
   hm  24. oct 2007        rev 1.4
       changed dst calculation because function dst was upgraded no error in DCF77 only a change in DST

   hm  12. nov 2007        rev 1.5
       changed time_offset from time to integer to allow for negative offset time zones

   hm  8. dec 2007     rev 1.6
       corrected an error in time_zone calculation

   hm 23. jan 2008     rev 1.7
       added sdt input which is used to initialize rtc and rtc1 during first cycle.

   hm 16. mar 2008     rev 1.8
       changed output weekday to wday and dst to ds for compatibility reasons

   hm  19. apr. 2008   rev 1.9
       added input dsi to allow to set daylight savings time when SDT is TRUE.
       added asynchronous SET input

   hm  7. oct. 2008    rev 1.10
       changed function weekday to day_of_week

   *)
END_FUNCTION_BLOCK

FUNCTION_BLOCK "HOLIDAY"   // FB28, SCL
TITLE = HOLIDAY
{ S7_Optimized_Access := 'FALSE' }
AUTHOR : hugo
FAMILY : TIDT
NAME : HOLIDAY
VERSION : 2.0
// holiday calculates if a given day is a holiday and displays the name of the holiday as string as well as a boolean flag to indicate a holiday.
// the holidays are specified in the country setup under global constants.
// a holiday can be of fixed date for example new years day on january 1st.
// a holiday can have a fixed offset from easter sunday as for most church holidays.
// a holiday can be a specific weekday before a fixed date, for example buss und bettag is the last wednesday before nov 23rd.
// with a simple f_use flag any specific holiday can be turned on or off if needed.
// 
// uses: LOCATION (DB5)
//       HOLIDAY_DATA (UDT9)
//       YEAR_OF_DATE (FC219)
//       EASTER (FC186)
//       SET_DATE (FC213)
//       LEAP_YEAR (FC194)
//       DAY_OF_WEEK (FC179)
//       DATE_ADD (FC176)
//       MONTH_OF_DATE (FC202)
//       DAY_OF_YEAR (FC180)
//       DATE_DINT (FC405)
//       LEAP_OF_DATE (FC193)
//       DAY_OF_MONTH (FC178)
   VAR_INPUT
      DATE_IN : Date;
      LANGU : Int;
      FRIDAY : Bool;
      SATURDAY : Bool;
      SUNDAY : Bool;
      SIZE : Int := 29;
   END_VAR
   VAR_OUTPUT
      Y : Bool;
      _NAME : String[30];
   END_VAR
   VAR_IN_OUT
      HOLIDAYS : Array[0..29] of "HOLIDAY_DATA";
   END_VAR
   VAR
      last_active : Date;
      ostern : Date;
      i : Int;
      jahr : Int;
      x_date : Date;
      lx : Int;
      wdx : Int;
   END_VAR
BEGIN


   (* for performance reasons only activate once a day *)
   IF #last_active = #DATE_IN THEN RETURN; END_IF;
   #last_active := #DATE_IN;

   (* determine language *)
   IF #LANGU = 0 THEN
     #lx := "LANGUAGE".DEFAULT;
   ELSE
     #lx := MIN(IN1:="LANGUAGE".LMAX,IN2:=#LANGU);
   END_IF;

   (* berechnung von ostern für das aktuelle jahr *)
   #jahr := "YEAR_OF_DATE"(#DATE_IN);
   #ostern := "EASTER"(#jahr);
   #wdx := "DAY_OF_WEEK"(#DATE_IN);
   #Y := FALSE;

   (* check for holidays *)
   FOR #i := 0 TO #SIZE DO
     #x_date := "SET_DATE"(YEAR:=#jahr, MONTH:=#HOLIDAYS[#i].MONTH , DAY:=#HOLIDAYS[#i].DAY);
     IF #HOLIDAYS[#i].USE = 1 AND #HOLIDAYS[#i].MONTH > 0 THEN
       (* check for fixed date holiday *)
       IF #x_date = #DATE_IN THEN
         #Y := TRUE;
         #_NAME := #HOLIDAYS[#i]BLKMOV_NAME;
         RETURN;
       END_IF;
     ELSIF #HOLIDAYS[#i].USE = 1 AND #HOLIDAYS[#i].MONTH = 0 THEN
       (* check for holiday in reference to easter *)
       IF "DATE_ADD"(IDATE:=#ostern, D:=#HOLIDAYS[#i].DAY ,W:=0,M:=0,Y:=0) = #DATE_IN THEN
         #Y := TRUE;
         #_NAME := #HOLIDAYS[#i]._NAME;
         RETURN;
       END_IF;
     ELSIF #HOLIDAYS[#i].USE < 0 THEN
       (* check for holiday on a weekday before date *)
       IF "DAY_OF_WEEK"(#DATE_IN) = ABS(#HOLIDAYS[#i].USE) AND #DATE_IN < #x_date AND #DATE_IN >= "DATE_ADD"(IDATE:=#x_date,D:=-7,W:=0,M:=0,Y:=0) THEN
         #Y := TRUE;
         #_NAME := #HOLIDAYS[#i]._NAME;
         RETURN;
       END_IF;
     END_IF;
   END_FOR;

   (* check array if today is weekend *)
   IF NOT #Y AND (#wdx = 5 AND #FRIDAY OR #wdx = 6 AND #SATURDAY OR #wdx = 7 AND #SUNDAY) THEN
     #Y := TRUE;
     #_NAME := "LANGUAGE".WEEKDAYSBLKMOV"LOCATION".LANGUAGE[#lx],#wdx];
   ELSE
     #_NAME := '';
   END_IF;


   (*
   Neujahrstag   1. Januar   •   •   •   •   •   •   •   •   •   •   •   •   •   •   •   •
   Heilige Drei Könige   6. Januar   •   •                         •     
   Karfreitag  Ostersonntag - 2d   •   •   •   •   •   •   •   •   •   •   •   •   •   •   •   •
   Ostersonntag  siehe Osterdatum        (•)                         
   Ostermontag   Ostersonntag + 1d   •   •   •   •   •   •   •   •   •   •   •   •   •   •   •   •
   Tag der Arbeit   1. Mai  •   •   •   •   •   •   •   •   •   •   •   •   •   •   •   •
   Christi Himmelfahrt   Ostersonntag + 39d  •   •   •   •   •   •   •   •   •   •   •   •   •   •   •   •
   Pfingstsonntag  Ostersonntag + 49d        (•)                         
   Pfingstmontag   Ostersonntag + 50d  •   •   •   •   •   •   •   •   •   •   •   •   •   •   •   •
   Fronleichnam  Ostersonntag + 60d  •   •           •       •   •   •   1)      2)
   Augsburger Friedensfest   8. August     (3)                             
   Mariä Himmelfahrt   15. August    (5)                     •         
   Tag der Deutschen Einheit   3. Oktober 6)   •   •   •   •   •   •   •   •   •   •   •   •   •   •   •   •
   Reformationstag   31. Oktober         •         •           •   •     •
   Allerheiligen   1. November   •   •                 •   •   •         
   Buß- und Bettag 4)  Mittwoch vor dem 23.11.       7                     •       
   1. Weihnachtstag  25. Dezember  •   •   •   •   •   •   •   •   •   •   •   •   •   •   •   •
   2. Weihnachtstag  26. Dezember  •   •   •   •   •   •   •   •   •   •   •   •   •   •   •   •
   *)



   (* revision history
   hm  27. feb. 2007 rev 1.1
     deleted unused variable init

   hm  31. oct. 2007 rev 1.2
     changed holiday definition from constant to input constant to allow easier changes by user without recompilation of the lib

   hm  24. nov. 2007 rev 1.3
     changes F_use of  Buß_und_Bettag to 0 because this is no official holiday

   hm  7. apr. 2008  rev 1.4
     improved performance

   hm  7. oct. 2008  rev 1.5
     changed code to use setup data from global constants
     changed length of output NAME from 20 to 30
     holiday will now also be indicated on a weekend
     changed function year to year_of_date
     changed function weekday to day_of_week

   hm  21. oct. 2008 rev 1.6
     using location constants

   hm  18. jan 2011  rev 2.0
     using user specified array for holidays

   *)
END_FUNCTION_BLOCK

FUNCTION_BLOCK "RTC_2"   // FB29, SCL
TITLE = RTC_2
{ S7_Optimized_Access := 'FALSE' }
AUTHOR : hugo
FAMILY : TIDT
NAME : RTC_2
VERSION : 1.4
// RTC_2 is a real time clock module which runs utc and generates local time from utc.
// daylight savings time can be enabled with den and an additional local time is generated with a delay of ofs im minutes.
// 
// uses: RTC_MS [FB30]
//       AD_DT_TM [FC1] 
//       T_PLC_MS [FC64] 
//       STIME [FB64],IDB_STIME [DB64] 
//       DST [FC183]
//       YEAR_OF_DATE [FC219] 
//       DT_DATE [FC6] 
//       DT_DINT [FC400] 
//       DT_TOD [FC8]
//       SET_DT [FC214] 
//       DINT_DT [FC399]
//       D_TOD_DT [FC3]
   VAR_INPUT
      SET : Bool;
      SDT : Date_And_Time;
      SMS : Int;
      DEN : Bool;
      OFS : Int;
   END_VAR
   VAR_OUTPUT
      _UDT : Date_And_Time;
      LDT : Date_And_Time;
      DSO : Bool;
      XMS : Int;
   END_VAR
   VAR
      RT : "RTC_MS";
   END_VAR
BEGIN


     (* call rtc *)
     #RT(SET := #SET, SDT := #SDT, SMS := #SMS);
     #_UDT := #RT.XDT;
     #XMS := #RT.XMS;

     (* check for daylight savings time and set dso output *)
     #DSO := "DST"(#_UDT) AND #DEN;

     (* calculate time offset and set ldt output *)
     #LDT := "DINT_DT"("DT_DINT"(#_UDT) + (#OFS + BOOL_TO_INT(#DSO)*60) * 60);


   (* revision history
   hm    20. jan. 2008  rev 1.0
     original version

   hm    20. feb. 2008  rev 1.1
     added Millisecond Set input

   hm    12. jun. 2008  rev 1.2
     improved performance

   hm    20. jan. 2011  rev 1.3
     changed offset to be in minutes

   hm    27. apr. 2011  rev 1.4
     fixed error with local time calculation

   *)
END_FUNCTION_BLOCK

FUNCTION_BLOCK "RTC_MS"   // FB30, SCL
TITLE = RTC_MS
{ S7_Optimized_Access := 'FALSE' }
AUTHOR : hugo
FAMILY : TIDT
NAME : RTC_MS
VERSION : 1.1
// RTC_MS is a real time clock module which can be set to SDT when set is TRUE and the outputs XDT and XT present the DateTime and TOD with a resolution of milliseconds.
// 
// uses: AD_DT_TM [FC1]
//       T_PLC_MS [FC64]
//       STIME [FB64],IDB_STIME [DB64]
   VAR_INPUT
      SET : Bool;
      SDT : Date_And_Time;
      SMS : Int;
   END_VAR
   VAR_OUTPUT
      XDT : Date_And_Time;
      XMS : Int;
   END_VAR
   VAR
      init : Bool;
      last : DWord;
      Tx : DWord;
   END_VAR
BEGIN


     #Tx := "T_PLC_MS"();
     IF #SET OR NOT #init THEN
       (* clock needs to be set when set is true or after power up *)
       #init := TRUE;
       #XDT := #SDT;
       #XMS := #SMS;
     ELSE
       #XMS := #XMS + DINT_TO_INT(DWORD_TO_DINT(#Tx) - DWORD_TO_DINT(#last));
       (* check if one second has expired *)
       IF #XMS > 999 THEN
         #XDT := #XDT T_ADD T#1s;
         #XMS := #XMS - 1000;
       END_IF;
     END_IF;
     #last := #Tx;


   (* revision history
   hm    20. jan. 2008 rev 1.0
     original version

   hm    20. feb. 2008 rev 1.1
     added Millisecond Set input
   *)
END_FUNCTION_BLOCK

FUNCTION_BLOCK "SUN_POS"   // FB31, SCL
TITLE = SUN_POS
{ S7_Optimized_Access := 'FALSE' }
AUTHOR : hugo
FAMILY : TIDT
NAME : SUNPOS
VERSION : 2.1
// this FUNCTION block calculates the sun position for a given date and time.
// the times are calculated in utc and have to be corrected for the given time zone.
// B is the angle from north and HR is the highth in degrees.
// 
// uses: DT_DATE [FC6]
//       DT_TOD [FC8]
//       MODR [FC97]
//       FLOOR2 [FC82] 
//       RAD [FC100]
//       DEG [FC72]
//       REFRACTION [FC206]
   VAR_INPUT
      latitude : Real;
      longitude : Real;
      utc : Date_And_Time;
   END_VAR
   VAR_OUTPUT
      "B" : Real;
      H : Real;
      HR : Real;
   END_VAR
   VAR
      g : Real;
      "a" : Real;
      d : Real;
      t1 : Real;
      n : Real;
      "e" : Real;
      c : Real;
      tau : Real;
      sin_d : Real;
      rlat : Real;
      sin_lat : Real;
      cos_lat : Real;
      cos_tau : Real;
      cos_d : Real;
   END_VAR
   VAR_TEMP
      temp_utc_DATE : Date;
      temp_utc_TOD : Time_Of_Day;
      temp : DInt;
   END_VAR
BEGIN


   (* n is the julian date and the number of days since 1.1.2000-12:00 midday *)
   (* be careful for step7 date startes 1.1.1990 instead of 1.1.1970 *)
   (* for step7 this line must change *)
   #temp_utc_DATE := T_CONV(IN := #utc); // DATE
   #temp_utc_TOD := T_CONV(IN := #utc); // TIME_OF_DAY

   #temp := (T_CONV(#temp_utc_DATE) + 7305) * 86400;  
   #temp := #temp + T_CONV(#temp_utc_TOD) / 1000;

   (* n is the julian date and the number of days since 1.1.2000-12:00 midday *)
   (* be careful for step7 date startes 1.1.1990 instead of 1.1.1970 *)
   (* for step7 this line must change *)
   #n := (DINT_TO_REAL(#temp) - 946728000) * 0.000011574074074074;
   #g := "MODR"(IN:=6.240040768 + 0.01720197 * #n, DIVI:="PI2_FB31");
   #d := "MODR"(IN:=4.89495042 + 0.017202792 * #n, DIVI:="PI2_FB31") + 0.033423055 * SIN(#g) + 0.000349066 * SIN(2.0*#g);
   #"e" := 0.409087723 - 0.000000006981317008 * #n;
   #cos_d := COS(#d);
   #sin_d := SIN(#d);
   #"a" := ATAN(COS(#"e") * #sin_d / #cos_d);
   IF #cos_d < 0.0 THEN #"a" := #"a" + "PI"; END_IF;
   #c := ASIN(SIN(#"e") * #sin_d);

   (* also here we must be very careful utc is from 1.1.1970 for step7 the formula must change *)
   #tau := "RAD"("MODR"(IN:=6.697376 + (#n - 0.25) * 0.0657098245037645 + DINT_TO_REAL(T_CONV(T_CONV(#utc))) * 0.0000002785383333, DIVI:=24.0) * 15.0 + #longitude) - #"a";
   #rlat := "RAD"(#latitude);
   #sin_lat := SIN(#rlat);
   #cos_lat := COS(#rlat);
   #cos_tau := COS(#tau);
   #t1 := #cos_tau * #sin_lat - TAN(#c) * #cos_lat;
   #"B" := ATAN(SIN(#tau) / #t1);
   IF #t1< 0.0 THEN #"B" := #"B" + "PI2_FB31"; ELSE #"B" := #"B" + "PI"; END_IF;
   #"B" := "DEG"("MODR"(IN:=#"B", DIVI:="PI2_FB31"));
   #H := "DEG"(ASIN(COS(#c) * #cos_tau * #cos_lat +SIN(#c) * #sin_lat));
   IF #H > 180.0 THEN #H := #H - 360.0; END_IF;
   (* consider refraction *)
   #HR := #H + "REFRACTION"(#H);


   (* revision history
   hm  1. feb 2007 rev 1.0
       original version

   hm  6. jan 2008 rev 1.1
       performance improvements

   hm  18. jan 2008    rev 1.2
       further performance improvements
       only calculate once every 10 seconds

   hm  16. mar. 2008   rev 1.3
       added type conversion to avoid warnings under codesys 3.0

   hm  30. jun. 2008   rev 1.4
       added type conversions to avoid warnings under codesys 3.0

   hm  18. oct. 2008   rev 1.5
       using math constants

   hm  17. dec. 2008   rev 1.6
       angles below horizon are displayed in negative degrees

   hm  27. feb. 2009   rev 2.0
       new code with better accuracy

   hm  7. mar. 2009    rev 2.1
       refraction is added after angle normalization
       deleted 10 second lockout
       added output for astronomical heigth h
   *)
END_FUNCTION_BLOCK

FUNCTION_BLOCK "SUN_TIME"   // FB32, SCL
TITLE = SUN_TIME
{ S7_Optimized_Access := 'FALSE' }
AUTHOR : hugo
FAMILY : TIDT
NAME : SUNTIME
VERSION : 1.7
// this FUNCTION block calculates the sun rise, sun set, sun offset at midday sun declination for a given date 
// for performance reasons the algorithm has been simplified and is accurate within a few minutes only 
// the times are calculated in utc and have to be corrected for the given time zone
// this correction is not done within sun_time because it would be a problem on days where dst is enabled or disabled
// 
// uses: SUN_MIDDAY (FC432)
//       DAY_OF_YEAR (FC180)
//       DATE_DINT (FC405)
//       HOUR_TO_TOD (FC190)
//       DEG (FC72)
//       MODR (FC97)
//       FLOOR2 (FC82)
//       HOUR_TO_TIME (FC189)
//       RAD (FC100)
   VAR_INPUT
      LATITUDE : Real;
      LONGITUDE : Real;
      UTC : Date;
      H : Real := -8.333333e-1;
   END_VAR
   VAR_OUTPUT
      MIDDAY : Time_Of_Day;
      SUN_RISE : Time_Of_Day;
      SUN_SET : Time_Of_Day;
      SUN_DECLINATION : Real;
   END_VAR
   VAR
      dk : Real;
      delta : Time;
      "b" : Real;
   END_VAR
BEGIN


   #"b" := #LATITUDE * 0.0174532925199433;
   #MIDDAY := "SUN_MIDDAY"(LON:=#LONGITUDE,UTC:=#UTC);
   #dk := 0.40954 * SIN(0.0172 * (INT_TO_REAL("DAY_OF_YEAR"(#UTC)) - 79.35));
   #SUN_DECLINATION := "DEG"(#dk);
   IF #SUN_DECLINATION > 180.0 THEN #SUN_DECLINATION := #SUN_DECLINATION - 360.0; END_IF;
   #SUN_DECLINATION := 90.0 - #LATITUDE + #SUN_DECLINATION;
   #delta := "HOUR_TO_TIME"(ACOS((SIN("RAD"(#H)) - SIN(#"b") * SIN(#dk)) / (COS(#"b") * COS(#dk))) * 3.819718632);
   #SUN_RISE := #MIDDAY - #delta;
   #SUN_SET := #MIDDAY + #delta;

   (* revision history

   rev 1.1 hm  20.1.2007
     deleted unused variables sun_riseR and sun_setR

   rev 1.2 hm 17.4.2007
     corrected error while sun:midday would not be corrected for longitude.

   rev 1.3 hm  6. jan 2008
     performance improvements

   rev 1.4 hm  17. jan 2008
     calculation is now only performed once a day

   hm  10. mar. 2009 rev 1.5
     improved performance
     calculation will be performed on every call to allow movong installations

   hm  26. jul 2009  rev 1.6
     fixed a problem with wrong midday calculation

   hm  25. jan. 2011 rev 1.7
     using function sun_midday
     corrected angle of sun_declination
     added input H
   *)
END_FUNCTION_BLOCK

FUNCTION_BLOCK "STIME"   // FB64, SCL
TITLE = STIME
{ S7_Optimized_Access := 'FALSE' }
AUTHOR : dalbi
FAMILY : MEASURE
NAME : STIME
VERSION : 1.4
// this function block makes sure that the timer of a siemens sps counts from 0 - 2^32-1.
   VAR_OUTPUT
      tx : DWord;
      at_tx AT tx : Array[0..31] of Bool;
   END_VAR
   VAR
      last_time : DWord;
      bit31 : Bool;
      init : Bool := TRUE;
   END_VAR
   VAR_TEMP
      TOP_SI : Struct
         EV_CLASS : Byte;
         EV_NUM : Byte;
         PRIORITY : Byte;
         NUM : Byte;
         TYP2_3 : Byte;
         TYP1 : Byte;
         ZI1 : Word;
         ZI2_3 : DWord;
      END_STRUCT;
      START_UP_SI : Struct
         EV_CLASS : Byte;
         EV_NUM : Byte;
         PRIORITY : Byte;
         NUM : Byte;
         TYP2_3 : Byte;
         TYP1 : Byte;
         ZI1 : Word;
         ZI2_3 : DWord;
      END_STRUCT;
      ERR : Int;
   END_VAR
BEGIN


   (* this FB is only necessary for siemens sps
   the siemens sps timer counts from 0 to 2^31-1 and starts at 0 sfter overrun.
   this means that the bit 31 (the highest bit ) will never be used and therefore
   a problem arises when t2 - t1 is checked.
   t2 - t1 is always valid also in an timer overrun situation where the time t1 is very high and t2 is very low.
   the result of the subtraction t2 - t1 however is still valid.
   this calculation does not work for soiemens because the highest bit is not used.

   this module stores the highest bit, changes the highest bit at every overrun occurence and stuffs ther highest bit in the output.
   the output is then used by t_plc_us and t_plc_ms.

   the correction needs and fb and not a function because the value of the highest bit has to be stored.

   do never use this function block in a codesys environment. the timer in codesys is correct and runs from 0 to 2^32-1
   *)

   (* read actual startup info *)
   (* OB1_SCAN_1  BYTE  -  B#16#01: Abschluss des Neustarts (Warmstarts)
                        -  B#16#02: Abschluss des Wiederanlaufs
                        -  B#16#03: Abschluss des freien Zyklus
                        -  B#16#04: Abschluss des Kaltstarts
                        -  B#16#05: Erster OB 1-Zyklus der neuen Master-CPU nach 
                                    Master-Reserve-Umschaltung und STOP des 
                                    bisherigen Masters *)

   #ERR := RD_SINFO (TOP_SI => #TOP_SI, START_UP_SI => #START_UP_SI);

   (* reset last_time on system startup *)
   IF #TOP_SI.EV_NUM = 1 OR #TOP_SI.EV_NUM = 2 OR #TOP_SI.EV_NUM = 4 OR NOT #init THEN 
       #last_time := 0;
       #bit31 := false;
       #init := true;
   END_IF;

   (* read the system timer *)
   #tx := DINT_TO_DWORD(T_CONV(TIME_TCK()));

   (* check for overrun *)
   IF DWORD_TO_DINT(#tx) < DWORD_TO_DINT(#last_time) THEN
       (* an overrun has occured, change the value of the highest bit *)
       #bit31 := NOT #bit31;
   END_IF;

   (* stuff the highest bit into the timer value *)
   #at_tx[7] := #bit31;

   (* remember the last system time for the next overrun check *)
   #last_time := #tx;


   (* revision history
   DA  14.9.2007 rev 1.0
     original version

   DA  24.2.2008 rev 1.1
     added self reset on system startup

   DA   2.5.2008 rev 1.2
     corect a problem running under OB35

   DA  12.3.2009 rev 1.3
     corect a problem run on different CPUs

   DA  22.12.2009 rev 1.4
     corect a problem on startup
   *)
END_FUNCTION_BLOCK

FUNCTION_BLOCK "EVENTS"   // FB254, SCL
TITLE = EVENTS
{ S7_Optimized_Access := 'FALSE' }
AUTHOR : hugo
FAMILY : TIDT
NAME : EVENTS
VERSION : 1.0
// event checks an array with a list of events and displays the event if today is one.
// 
// uses: DAY_OF_DATE (FC177)
//       YEAR_OF_DATE (FC219)
//       SET_DATE (FC213)
//       LEAP_YEAR (FC194)
//       HOLIDAY_DATA (UDT9)
   VAR_INPUT
      DATE_IN : Date;
      ENA : Bool;
   END_VAR
   VAR_OUTPUT
      Y : Bool;
      _NAME : String[30];
   END_VAR
   VAR_IN_OUT
      ELIST : Array[0..49] of "HOLIDAY_DATA";
   END_VAR
   VAR
      i : Int;
      last_active : Date;
      size : Int := 49;
      day_in : DInt;
      cyr : Int;
      lday : DInt;
      check : "HOLIDAY_DATA";
      y_int : Bool;
      name_int : String[30];
   END_VAR
BEGIN


   (* for performance reasons only activate once a day *)
   IF #last_active <> #DATE_IN THEN
     #last_active := #DATE_IN;
     #y_int := FALSE;
     #name_int := '';
     #day_in := "DAY_OF_DATE"(#DATE_IN);
     #cyr := "YEAR_OF_DATE"(#DATE_IN);

     (* search list for events *)
     FOR #i := 0 TO #size DO
       #check := #ELIST[#i];
       #lday := "DAY_OF_DATE"("SET_DATE"(YEAR:=#cyr,MONTH:=#check.MONTH,DAY:=#check.DAY));
       IF #day_in >= #lday AND #day_in <= #lday + #check.USE - 1 THEN
         #y_int := TRUE;
         #name_int BLKMOV #check._NAME;
         EXIT;
       END_IF;
     END_FOR;
   END_IF;

   IF #ENA THEN
     #Y := #y_int;
     #_NAME BLKMOV #name_int;
   ELSE
     #Y := FALSE;
     #_NAME := '';
   END_IF;


   (* revision history
   hm  18. jan. 2011 rev 1.0
     new module

   *)
END_FUNCTION_BLOCK

FUNCTION "T_PLC_MS" : DWord   // FC64, SCL
TITLE = T_PLC_MS
{ S7_Optimized_Access := 'FALSE' }
AUTHOR : hugo
FAMILY : MEASURE
NAME : T_PLC_MS
VERSION : 1.2
// T_PLC_MS reads the internal PLC timer and return the time, it has the advantage to be able to set a debug mode 
// and speed up the counter to test the plc timer overrun which occurs every 50 days respectively 25 days at siemens S7
// this routine also allows to correct the behavior of s7 where the internal plc counter will not count all 32 bits.
// 
// uses: STIME [FB64],IDB_STIME [DB64]
BEGIN


   "IDB_STIME"(); 
   #T_PLC_MS := "IDB_STIME".tx; 
   (* hier muss die korrektur für step7 stattfinden
   plctime muss den vollen wertebereich von time ausnutzen:
   wenn bei step7 time -24tage bis plus 24 tage ist dann muss der timer auch beim überlauf auf -24tage springen 
   und auf keinen fall auf 0 !!!!
   für siemens muss ein weiterer fb im main eingebunden werden der sicherstellt das alle 32 bits durchgezählt werden.
   es kann nur ein fb sein den er muss sich das oberste (32te) bit merken.
   oder etwa spring s7 bei überlauf auf -24 tage????? dann wäre keine korrektur nötig.
   *)
   IF "debug" THEN
       #T_PLC_MS := DINT_TO_DWORD((DWORD_TO_DINT(SHL(IN:=#T_PLC_MS,N:="N") OR SHL(IN:=DWORD#1,N:="N"))-1) + DWORD_TO_DINT("offset_1"));
   END_IF;


   (* revision history
   hm  14.9.2007   rev 1.0
       original version

   hm  12. nov 2007    rev 1.1
       added temporaray variable tx because some compilers could not handle time() as an argument

   hm  16. nov. 2008   rev 1.2
       initialized constants with 0 for compatibility reasons
   *)
END_FUNCTION

FUNCTION "DEG" : Real   // FC72, SCL
TITLE = DEG
{ S7_Optimized_Access := 'FALSE' }
AUTHOR : hugo
FAMILY : MATH
NAME : DEG
VERSION : 1.2
// this function converts degrees into Radiant
// 
// uses: MODR [FC97]
//       FLOOR2 [FC82]
   VAR_INPUT
      rad : Real;
   END_VAR
BEGIN


   #DEG := "MODR"(IN:=57.29577951308232 * #rad,DIVI:=360.0);


   (* revision history
   hm  4. aug 2006 rev 1.0
       original version

   hm 16. oct 2007 rev 1.1
       added modr statement which prohibits deg to become bigger than 360

   hm  10. mar. 2009   rev 1.2
       real constants updated to new systax using dot
   *)
END_FUNCTION

FUNCTION "EVEN" : Bool   // FC76, SCL
TITLE = EVEN
{ S7_Optimized_Access := 'FALSE' }
AUTHOR : hugo
FAMILY : MATH
NAME : EVEN
VERSION : 1.2
// this function chacks an input for even value
// the output is true if the input is even.
   VAR_INPUT
      in : DInt;
   END_VAR
   VAR_TEMP
      tIN : DInt;
      _IN AT tIN : Array[0..31] of Bool;
   END_VAR
BEGIN


   #tIN := #in;
   #EVEN := NOT #_IN[24]; //EVEN := NOT in.0;

   (* revision history
   hm  1. oct 2006 rev 1.0
     ORIGINAL VERSION

   hm  01.12.2007  rev 1.1
     changed code for improved performance

   hm  21. mar. 2008 rev 1.2
     changed type of input IN from INT to DINT
   *)
END_FUNCTION

FUNCTION "FLOOR2" : DInt   // FC82, SCL
TITLE = FLOOR2
{ S7_Optimized_Access := 'FALSE' }
AUTHOR : hugo
FAMILY : MATH
NAME : FLOOR2
VERSION : 1.1
// This is a rounding function which returns the biggest possible integer which is less or equal to X.
// floor2(3.14) = 3
// floor2(-3.14) = -4
   VAR_INPUT
      X : Real;
   END_VAR
BEGIN


   #FLOOR2 := REAL_TO_DINT(#X);
   IF DINT_TO_REAL(#FLOOR2) > #X THEN
     #FLOOR2 := #FLOOR2 - 1;
   END_IF;

   (* revision history
   hm  21. mar. 2008   rev 1.0
       originlal version

   hm  4. apr. 2008    rev 1.1
       added type conversion to avoid warnings under codesys 3.0
   *)
END_FUNCTION

FUNCTION "MODR" : Real   // FC97, SCL
TITLE = MODR
{ S7_Optimized_Access := 'FALSE' }
AUTHOR : hugo
FAMILY : MATH
NAME : MODR
VERSION : 1.5
// this is a modulo funtion for real numbers
// modr(5.5,2.5) = 0.5
// 
// uses: FLOOR2 [FC82]
   VAR_INPUT
      IN : Real;
      DIVI : Real;
   END_VAR
BEGIN


   IF #DIVI = 0.0 THEN
       #MODR := 0.0;
   ELSE
       #MODR := #IN - DINT_TO_REAL("FLOOR2"(#IN / #DIVI)) * #DIVI;
   END_IF;


   (* revision history

   hm  4. aug.2006     rev 1.0

   hm  28. jan.2007   rev 1.1
       modr(x,0) will deliver the result 0

   hm  21. mar 2008    rev 1.2
       use D_trunc for compatibility reasons

   hm  4. apr. 2008    rev 1.3
       added type conversion to avoid warnings under codesys 3.0

   hm  31. oct. 2008   rev 1.4
       changed algorithm to the more common version using floor instead of TRUNC

   hm  10. mar. 2009   rev 1.5
       real constants updated to new systax using dot

   *)
END_FUNCTION

FUNCTION "RAD" : Real   // FC100, SCL
TITLE = RAD
{ S7_Optimized_Access := 'FALSE' }
AUTHOR : hugo
FAMILY : MATH
NAME : RAD
VERSION : 1.2
// this function converts Radiant to degrees
// 
// uses: MODR [FC97]
//       FLOOR2 [FC82]
   VAR_INPUT
      deg : Real;
   END_VAR
BEGIN


   #RAD := "MODR"(IN:=0.0174532925199433 * #deg,DIVI:="PI2");

   (*  Enfällt da der Zugriff auf Datenbaustein länger dauert
       RAD := MODR(0.0174532925199433 * DEG, math.PI2);
   *)

   (* revision history
   hm  4. aug 2006     rev 1.0
       original version

   hm  16. oct 2007    rev 1.1
       added modr statement which prohibits rad to become bigger than 2PI

   hm  18. oct 2008    rev 1.2
       using math constants

   *)
END_FUNCTION

FUNCTION "DATE_ADD" : Date   // FC176, SCL
TITLE = DATE_ADD
{ S7_Optimized_Access := 'FALSE' }
AUTHOR : hugo
FAMILY : TIDT
NAME : DTADD
VERSION : 1.8
// date_add adds days, weeks, month or years to a date.
// negative inputs are allowed for subtraction.
// 
// uses: LEAP_YEAR [FC194] 
//       SET_DATE [FC213]
//       DATE_DINT [FC405]
//       LEAP_OF_DATE [FC193] 
//       DAY_OF_YEAR [FC180] 
//       DAY_OF_MONTH [FC178]
//       MONTH_OF_DATE [FC202]
//       YEAR_OF_DATE [FC219]
   VAR_INPUT
      IDATE : Date;
      D : Int;
      W : Int;
      "M" : Int;
      Y : Int;
   END_VAR
   VAR_TEMP
      mo : Int;
      yr : Int;
      dm : Int;
   END_VAR
BEGIN


   #DATE_ADD := T_CONV(T_CONV(#IDATE) + INT_TO_DINT(#D) + 7 * INT_TO_DINT(#W));
   #yr := #Y + "YEAR_OF_DATE"(#DATE_ADD);
   #mo := #"M" + "MONTH_OF_DATE"(#DATE_ADD);
   #dm := "DAY_OF_MONTH"(#DATE_ADD);
   WHILE #mo > 12 DO
     #mo := #mo - 12;
     #yr := #yr + 1;
   END_WHILE;
   WHILE #mo < 1 DO
     #mo := #mo + 12;
     #yr := #yr - 1;
   END_WHILE;
   #DATE_ADD := "SET_DATE"(YEAR:=#yr,MONTH:=#mo,DAY:=#dm);


   (* revision history

   hm 27.12.2006 rev 1.0
     nrw module

   hm 12.4.2007    rev 1.1
     corrected an error while date would be incorrect when year  = 0

   hm  1.11.2007   rev 1.2
     added int_to_dword stetements to avoid possible overrun with möller ecp4

   hm  22. mar. 2008 rev 1.3
     fixed some bugs when month was negative

   hm  7. oct. 2008  rev 1.4
     changed function year to year_of_date
     changed function month to month_of_date

   hm  29. mar. 2009 rev 1.5
     improved performance

   hm  27. jan. 2011 rev 1.6
     faster code

   hm  2. feb. 2011    rev 1.7
     fixed an error, weeks not calculated

   hm  22. mar. 2011 rev 1.8
     fixed an error in formula
   *)
END_FUNCTION

FUNCTION "DAY_OF_DATE" : DInt   // FC177, SCL
TITLE = DAY_OF_DATE
{ S7_Optimized_Access := 'FALSE' }
AUTHOR : oscat
FAMILY : TIDT
NAME : DAYDT
VERSION : 1.3
// DAY_OF_DATE returns the days since 1.1.1970
   VAR_INPUT
      idate : Date;
   END_VAR
   VAR_TEMP
      tDate : DInt;
   END_VAR
BEGIN


   (* adjust step7 day by 7305 days because step7 date format starts at 1.1.1990  *)
   #DAY_OF_DATE := T_CONV(#idate) + 7305; // 86400 sec format

   (*
   day_of_date := DWORD_TO_DINT(DATE_TO_DWORD(idate) / 86400);
   *)

   (* revision history
   hm      16.9.2007       rev 1.0
       original version

   hm      1. okt 2007     rev 1.1
       added step7 compatibility

   hm      22. mar. 2008   rev 1.2
       changed output from int to Dint because the total date range is 49710 days

   hm      7. apr. 2008    rev 1.3
       deleted unused step7 code

   *)
END_FUNCTION

FUNCTION "DAY_OF_MONTH" : Int   // FC178, SCL
TITLE = DAY_OF_MONTH
{ S7_Optimized_Access := 'FALSE' }
AUTHOR : hugo
FAMILY : TIDT
NAME : DAYOMON
VERSION : 2.1
// returns the day OF month from any DATE
// 
// uses: DAY_OF_YEAR [FC180]
//       YEAR_BEGIN [FC217] 
//       YEAR_OF_DATE [FC219] 
//       LEAP_OF_DATE [FC193]
//       LEAP_YEAR [FC194]
   VAR_INPUT
      IDATE : Date;
   END_VAR
   VAR_TEMP
      leap : Int;
   END_VAR
BEGIN


   (* calculate the day in the year *)
   #DAY_OF_MONTH := "DAY_OF_YEAR"(#IDATE);
   (* leap will be set to one for a leap year *)
   #leap := BOOL_TO_INT("LEAP_OF_DATE"(#IDATE));
   (* if leap year deduct one from the days of the year *)
   #DAY_OF_MONTH := #DAY_OF_MONTH - #leap;
   (* search if we are in month december to march ? *)
   IF #DAY_OF_MONTH > "MTH_OFS9" THEN
       IF #DAY_OF_MONTH > "MTH_OFS11" THEN
           IF #DAY_OF_MONTH > "MTH_OFS12" THEN
               #DAY_OF_MONTH := #DAY_OF_MONTH - "MTH_OFS12";
           ELSE
               #DAY_OF_MONTH := #DAY_OF_MONTH - "MTH_OFS11";
           END_IF;
       ELSE
           IF #DAY_OF_MONTH > "MTH_OFS10" THEN
               #DAY_OF_MONTH := #DAY_OF_MONTH - "MTH_OFS10";
           ELSE
               #DAY_OF_MONTH := #DAY_OF_MONTH - "MTH_OFS9";
           END_IF;
       END_IF;
   ELSIF #DAY_OF_MONTH > "MTH_OFS5" THEN
       IF #DAY_OF_MONTH > "MTH_OFS7" THEN
           IF #DAY_OF_MONTH > "MTH_OFS8" THEN
               #DAY_OF_MONTH := #DAY_OF_MONTH - "MTH_OFS8";
           ELSE
               #DAY_OF_MONTH := #DAY_OF_MONTH - "MTH_OFS7";
           END_IF;
       ELSE
           IF #DAY_OF_MONTH > "MTH_OFS6" THEN
               #DAY_OF_MONTH := #DAY_OF_MONTH - "MTH_OFS6";
           ELSE
               #DAY_OF_MONTH := #DAY_OF_MONTH - "MTH_OFS5";
           END_IF;
       END_IF;
   ELSIF #DAY_OF_MONTH > "MTH_OFS3" THEN
       IF #DAY_OF_MONTH > "MTH_OFS4" THEN
           #DAY_OF_MONTH := #DAY_OF_MONTH - "MTH_OFS4";
       ELSE
           #DAY_OF_MONTH := #DAY_OF_MONTH - "MTH_OFS3";
       END_IF;
   ELSE
       (* since now we must be in february or january we need to add leap again *)
       #DAY_OF_MONTH := #DAY_OF_MONTH + #leap;
       IF #DAY_OF_MONTH > "MTH_OFS2" THEN #DAY_OF_MONTH := #DAY_OF_MONTH - "MTH_OFS2"; END_IF;
       (* since nothing was true before, day_of_month must already be good *)
   END_IF;


   (*
   Revision history

   hm 22.1.2007        rev 1.1
       deleted unused variable day_in_year and day_in_year_begin

   hm  1. okt 2007 rev 1.2
       changed code to use day_of_year and leap_of_date
       added compatibility to STEP7

   hm  8. oct 2007 rev 1.3
       deleted unused variable yr

   hm  8. jan 2008 rev 1.4
       improved performance

   hm  25. oct. 2008   rev 2.0
       new code using setup constants

   hm  10. mar. 2009   rev 2.1
       removed nested comments

   *)
END_FUNCTION

FUNCTION "DAY_OF_WEEK" : Int   // FC179, SCL
TITLE = DAY_OF_WEEK
{ S7_Optimized_Access := 'FALSE' }
AUTHOR : hugo
FAMILY : TIDT
NAME : DWEEK
VERSION : 1.4
// calculates the weekday of a week according to ISO8601   
// monday = 1 ..... sunday = 7
   VAR_INPUT
      IDATE : Date;
   END_VAR
BEGIN


     #DAY_OF_WEEK := DINT_TO_INT((T_CONV(#IDATE)+7308) MOD 7)+1;

   (* 
   weekday := DWORD_TO_INT((DATE_TO_DWORD(idate)/86400+3) MOD 7) + 1;
   *)


   (* revision history
   hm  21.8.06         rev 1.1
       corrected a miscalculation

   hm  23.12.2007      rev 1.2
       correction for step7

   hm  7. apr. 2008    rev 1.3
       deleted unused step7 code

   hm  7. oct. 2008    rev 1.4
       changed name of function from weekday to day_of_week

   *)
END_FUNCTION

FUNCTION "DAY_OF_YEAR" : Int   // FC180, SCL
TITLE = DAY_OF_YEAR
{ S7_Optimized_Access := 'FALSE' }
AUTHOR : hugo
FAMILY : TIDT
NAME : DAYOYEAR
VERSION : 1.4
// calculates the day of the year
// 
// uses: DATE_DINT [FC405]
   VAR_INPUT
      idate : Date;
   END_VAR
BEGIN


   #DAY_OF_YEAR := DINT_TO_INT(("DATE_DINT"(#idate) / 86400) MOD 1461);
   IF #DAY_OF_YEAR > 729 THEN
     IF #DAY_OF_YEAR > 1095 THEN #DAY_OF_YEAR := #DAY_OF_YEAR - 1095; ELSE #DAY_OF_YEAR := #DAY_OF_YEAR - 729; END_IF;
   ELSIF #DAY_OF_YEAR > 364 THEN
     #DAY_OF_YEAR := #DAY_OF_YEAR - 364;
   ELSE
     #DAY_OF_YEAR := #DAY_OF_YEAR + 1;
   END_IF;

   //  day_of_year := DINT_TO_INT((DATE_TO_DINT(idate) - DATE_TO_DINT(year_begin(year_of_date(idate))))) + 1;

   (*
   DAY_OF_YEAR := DWORD_TO_INT((DATE_TO_DWORD(idate) - DATE_TO_DWORD(YEAR_BEGIN(YEAR_OF_DATE(idate)))) / 86400) + 1;
   *)


   (* revivision history
   hm  4. aug. 2007    rev 1.0
     original version

   hm  1. oct. 2007    rev 1.1
     added compatibility to STEP7

   hm  4. jan. 2008    rev 1.2
     changed code for better performance

   hm  7. oct. 2008    rev 1.3
     changed name of function year to year_of_date

   hm  28. jan. 2011 rev 1.4
     improved code
   *)
END_FUNCTION

FUNCTION "DAY_TO_TIME" : Time   // FC181, SCL
TITLE = DAY_TO_TIME
{ S7_Optimized_Access := 'FALSE' }
AUTHOR : hugo
FAMILY : TIDT
NAME : DAY2TI
VERSION : 1.1
// converts an amount of days in real to time
   VAR_INPUT
      IN : Real;
   END_VAR
BEGIN


   #DAY_TO_TIME := T_CONV(REAL_TO_DINT(#IN * 86400000));


   (* revision history
   hm  4. aug. 2006    rev 1.0
       original release

   hm  24. feb. 2009   rev 1.1
       renamed input to IN
   *)
END_FUNCTION

FUNCTION "DAYS_DELTA" : DInt   // FC182, SCL
TITLE = DAYS_DELTA
{ S7_Optimized_Access := 'FALSE' }
AUTHOR : hugo
FAMILY : TIDT
NAME : DAYDELT
VERSION : 1.3
// days_delta calculates the days between two dates. the days are calculated date_2 - date_1
   VAR_INPUT
      date_1 : Date;
      date_2 : Date;
   END_VAR
BEGIN


     IF T_CONV(#date_1) > T_CONV(#date_2) THEN
       #DAYS_DELTA := - (T_CONV(#date_1) - T_CONV(#date_2));
     ELSE
       #DAYS_DELTA := T_CONV(#date_2) - T_CONV(#date_1);
     END_IF;

     //days_delta := day_of_date(date_2) - day_of_date(date_1);

   (* revision history
   hm  27. dec 2006  rev 1.0
     original version

   hm  16.9.2007   rev 1.1
     coorected an error in formula and changed algorithm to show positive and negative delta

   hm  22. mar. 2008 rev 1.2
     changed output from int to dint because the total date range is 49710 days

   hm  25. jan. 2011 rev 1.3
     improved performance
   *)
END_FUNCTION

FUNCTION "DST" : Bool   // FC183, SCL
TITLE = DST
{ S7_Optimized_Access := 'FALSE' }
AUTHOR : hugo
FAMILY : TIDT
NAME : DST
VERSION : 1.5
// this functions returns TRUE IF dst TIME is active 
// the FUNCTION calculates automatically for any year betweek 1970 AND 2099 
// wheather daylight savings is on OR off 
// the summertime calculation is done according to european standards.
// dst will become TRUE AT 01:00 utc in the morning FOR the respective days 
// AND it will become FALSE after daylight savings TIME is switched back end OF october at 01:00 utc
// 
// uses: YEAR_OF_DATE [FC219]
//       DT_DATE [FC6]
//       DT_DINT [FC400]
//       DT_TOD [FC8] 
//       SET_DT [FC214]
   VAR_INPUT
      UTC : Date_And_Time;
   END_VAR
   VAR_TEMP
      temp_utc : Date_And_Time;
      yr : Int;
      yr4 : DInt;
      ltc : DInt;
      idate : DInt;
   END_VAR
BEGIN


   #temp_utc := #UTC;

   #yr := "YEAR_OF_DATE"(T_CONV(#temp_utc));
   #ltc := "DT_DINT"(#temp_utc);
   #idate := "DT_DINT"("SET_DT"(year:=#yr,month:=3,day:=31,hour:=1,minute:=0,second:=0));
   #yr4 := DWORD_TO_DINT(SHR(IN:=DINT_TO_DWORD(5*INT_TO_DINT(#yr)),N:=2)) + 1;
   #DST := (#idate - ((#yr4 + 3) MOD 7) * 86400 <= #ltc) AND (#idate + (214 - (#yr4) MOD 7) * 86400 > #ltc);


   (*
   Equation used TO calculate the beginning OF European Summer TIME:
   Sunday (31 - (5*y/4 + 4) mod 7) March at 01.00 UTC
   (valid through 2099, courtesy of Robert H. van Gent, EC).

   European Summer Time ends (clocks go back) at 01.00 UTC on

       * 29 October 2006
       * 28 October 2007
       * 26 October 2008

   Equation used to calculate the end of European Summer Time:
   Sunday (31 - (5*y/4 + 1) mod 7) October at 01.00 UTC
   (validity AND credits as above).

   *)



   (* revision history
   hm  4. aug 2006 rev 1.0
     original version

   hm  24. okt 2007  rev 1.1
     deleted time_zone_offset input because dst is generally at 01:00 utc and not mesz
     uk starts 01:00 utc and also greece

   hm  1. dec 2007 rev 1.2
     changed code to improve performance

   hm  16. mar. 2008 rev 1.3
     added type conversion to avoid warnings under codesys 3.0
     code improvement for better performance

   hm  7. oct. 2008  rev 1.4
     changed name of function year to year_of_date

   hm  24. jan. 2011 rev 1.5
     improved performance
   *)
END_FUNCTION

FUNCTION "DT2_TO_SDT" : "SDT"   // FC184, SCL
TITLE = DT2_TO_SDT
{ S7_Optimized_Access := 'FALSE' }
AUTHOR : hugo
FAMILY : TIDT
NAME : DT2SDT
VERSION : 1.0
// converts date and time of day to Structured date time (SDT)
// 
// uses: SDT [UDT12]
//       D_TOD_DT [FC3]
   VAR_INPUT
      _DI : Date;
      TI : Time_Of_Day;
   END_VAR
   VAR_TEMP
      Year : Int;
      tMS : Word;
      tDTI : Date_And_Time;
      _DTI AT tDTI : Struct
         Year : Byte;
         Month : Byte;
         Day : Byte;
         Hour : Byte;
         Minute : Byte;
         Second : Byte;
         ms : Byte;
         wday_ms : Byte;
      END_STRUCT;
      tDT2_TO_SDT : "SDT";
   END_VAR
BEGIN


   #tDTI := T_COMBINE(IN1:=#_DI,IN2:=#TI);

   #Year := BCD16_TO_INT(#_DTI.Year);
   IF #Year >= 90 THEN 
       #tDT2_TO_SDT.YEAR := #Year + 1900; 
   ELSE 
       #tDT2_TO_SDT.YEAR := #Year + 2000; 
   END_IF;
   #tDT2_TO_SDT.MONTH := BCD16_TO_INT(#_DTI.Month);
   #tDT2_TO_SDT.DAY := BCD16_TO_INT(#_DTI.Day);
   #tDT2_TO_SDT.HOUR := BCD16_TO_INT(#_DTI.Hour);
   #tDT2_TO_SDT.MINUTE := BCD16_TO_INT(#_DTI.Minute);
   #tDT2_TO_SDT.SECOND := BCD16_TO_INT(#_DTI.Second);
   #tMS := SHL(IN:=BYTE_TO_WORD(#_DTI.ms),N:=4);
   #tMS := #tMS OR SHR(IN:=BYTE_TO_WORD(#_DTI.wday_ms),N:=4);
   #tDT2_TO_SDT.MS := BCD16_TO_INT(#tMS);
   #tDT2_TO_SDT.WEEKDAY := BCD16_TO_INT(SHR(IN:=SHL(IN:=#_DTI.wday_ms,N:=4),N:=4));

   #DT2_TO_SDT := #tDT2_TO_SDT;

   (* Original
   DT2_TO_SDT.YEAR := YEAR_OF_DATE(di);
   DT2_TO_SDT.MONTH := MONTH_OF_DATE(di);
   DT2_TO_SDT.DAY := DAY_OF_MONTH(di);
   DT2_TO_SDT.WEEKDAY := DAY_OF_WEEK(di);
   DT2_TO_SDT.MS := DWORD_TO_INT(TOD_TO_DWORD(ti) MOD 1000);
   DT2_TO_SDT.SECOND := DWORD_TO_INT((TOD_TO_DWORD(ti) / 1000) MOD 60);
   DT2_TO_SDT.MINUTE := DWORD_TO_INT((TOD_TO_DWORD(ti) / 60000) MOD 60);
   DT2_TO_SDT.HOUR := DWORD_TO_INT(TOD_TO_DWORD(ti) / 3600000);
   *)

   (* revision history

   hm 18. oct. 2008    rev 1.0
       original version

   *)
END_FUNCTION

FUNCTION "DT_TO_SDT" : "SDT"   // FC185, SCL
TITLE = DT_TO_SDT
{ S7_Optimized_Access := 'FALSE' }
AUTHOR : hugo
FAMILY : TIDT
NAME : DTSDT
VERSION : 1.0
// converts date_time to Structured date time (SDT)
// 
// uses: SDT [UDT12]
   VAR_INPUT
      DTI : Date_And_Time;
      _DTI AT DTI : Struct
         Year : Byte;
         Month : Byte;
         Day : Byte;
         Hour : Byte;
         Minute : Byte;
         Second : Byte;
         ms : Byte;
         wday_ms : Byte;
      END_STRUCT;
   END_VAR
   VAR_TEMP
      Year : Int;
      tMS : Word;
      tDT_TO_SDT : "SDT";
   END_VAR
BEGIN


   #Year := BCD16_TO_INT(#_DTI.Year);
   IF #Year >= 90 THEN 
       #tDT_TO_SDT.YEAR := #Year + 1900; 
   ELSE 
       #tDT_TO_SDT.YEAR := #Year + 2000; 
   END_IF;
   #tDT_TO_SDT.MONTH := BCD16_TO_INT(#_DTI.Month);
   #tDT_TO_SDT.DAY := BCD16_TO_INT(#_DTI.Day);
   #tDT_TO_SDT.HOUR := BCD16_TO_INT(#_DTI.Hour);
   #tDT_TO_SDT.MINUTE := BCD16_TO_INT(#_DTI.Minute);
   #tDT_TO_SDT.SECOND := BCD16_TO_INT(#_DTI.Second);
   #tMS := SHL(IN:=BYTE_TO_WORD(#_DTI.ms),N:=4);
   #tMS := #tMS OR SHR(IN:=BYTE_TO_WORD(#_DTI.wday_ms),N:=4);
   #tDT_TO_SDT.MS := BCD16_TO_INT(#tMS);
   #tDT_TO_SDT.WEEKDAY := BCD16_TO_INT(SHR(IN:=SHL(IN:=#_DTI.wday_ms,N:=4),N:=4));

   #DT_TO_SDT := #tDT_TO_SDT;


   (* revision history

   hm 18. oct. 2008    rev 1.0
       original version

   *)
END_FUNCTION

FUNCTION "EASTER" : Date   // FC186, SCL
TITLE = EASTER
{ S7_Optimized_Access := 'FALSE' }
AUTHOR : hugo
FAMILY : TIDT
NAME : EASTER
VERSION : 1.3
// easter calculates the day of easter sunday for a given year.
// most other catholic holidays are calculated in reference to easter sunday.
// 
// uses: SET_DATE [FC213]
//       LEAP_YEAR [FC194]
   VAR_INPUT
      year : Int;
   END_VAR
   VAR_TEMP
      "b" : Int;
      c : Int;
      oday : Int;
      omon : Int;
   END_VAR
BEGIN


   #"b" := (204 - 11 * (#year MOD 19)) MOD 30;
   IF #"b" > 27 THEN #"b" := #"b" - 1; END_IF;
   #c := (#year + WORD_TO_INT(SHR(IN:=INT_TO_WORD(#year),N:=2)) + #"b" - 13) MOD 7;
   #oday := 28 + #"b" - #c;
   IF #oday > 33 THEN
       #EASTER := "SET_DATE"(YEAR:=#year,MONTH:=4,DAY:=#oday - 31);
   ELSE
       #EASTER := "SET_DATE"(YEAR:=#year,MONTH:=3,DAY:=#oday);
   END_IF;

   (* alternativer algorithmus ueber das pasah fest
   execution time roughly 200us
   Der sog. Passah-Vollmond wird berechnet, in dem das Jahr durch 19 ge-
   teilt wird und der Rest mit der folgenden Tabelle verglichen wird:

       0: Apr 14       5: Apr 18      10: Mrz 25      15: Mrz 30
       1: Apr 03       6: Apr 08      11: Apr 13      16: Apr 17
       2: Mrz 23       7: Mrz 28      12: Apr 02      17: Apr 07
       3: Apr 11       8: Apr 16      13: Mrz 22      18: Mrz 27
       4: Mrz 31       9: Apr 05      14: Apr 10

   Faellt dieses Datum auf einen Sonntag, ist Ostern der naechste Sonntag!

   Beispiel: 1992 MOD 19 = 16, daraus folgt 17.04., der naechste Sonntag
             ist dann der 19. April (Ostersonntag)
   *)


   (* this algorithm is 180 us
   a := year MOD 19;
   b := year / 100;
   c := year MOD 100;
   d := b / 4;
   e := b MOD 4;
   f := (b + 8) / 25;
   g := (b - f + 1) / 3;
   h := (19 * a + b - d -g + 15) MOD 30;
   i := C / 4;
   k := c MOD 4;
   l := (32 + 2*e + 2*i - h - k) MOD 7;
   m := (a + 11 * h + 22 * l) / 451;
   x := h + l - 7 * m + 114;
   n := X / 31;
   o := x MOD 31 + 1;

   easter := set_Date(year,n,o);
   *)
   (*
   Im Magazin "Nature" vom 20. April 1876 veröffentlichte ein anonymer Autor eine Tabelle mit Regeln zur Berechnung des (Gregorianischen) Ostersonntages des Jahres J. In Formeln ausgedrückt erhält man das Folgende:
   a   =   J mod 19
   b   =   int(J / 100)
   c   =   J mod 100
   d   =   int(b / 4)
   e   =   b mod 4
   f   =   int((b + 8) / 25)
   g   =   int((b - f + 1) / 3
   h   =   (19 · a + b - d - g + 15) mod 30
   i   =   int(c / 4)
   k   =   c mod 4
   l   =   (32 + 2 · e + 2 · i - h - k) mod 7
   m   =   int((a + 11 · h + 22 · l) / 451)
   n   =   int((h + l - 7 · m + 114) / 31)
   o   =   (h + l - 7 · m + 114) mod 31

   n ist hierbei die Nummer des Monats, o + 1 die Nummer des Tages auf welchen der Ostersonntag im Jahr J fällt. Dieser Algorithmus kommt ohne Hilfszahlen aus.

   *)

   (* revision history
   hm  27. dec 2006    rev 1.0
       original version

   hm  15. dec 2007    rev 1.1
       modified code for better performance

   hm  3. feb 2008     rev 1.2
       modified code for better performance

   hm  7. apr. 2008    rev 1.3
       improved performance
   *)
END_FUNCTION

FUNCTION "HOUR" : Int   // FC187, SCL
TITLE = HOUR
{ S7_Optimized_Access := 'FALSE' }
AUTHOR : hugo
FAMILY : TIDT
NAME : HOUR
VERSION : 1.1
// extracts the hour of a Time_of_day
   VAR_INPUT
      itod : Time_Of_Day;
   END_VAR
BEGIN


     #HOUR := DINT_TO_INT(T_CONV(#itod)/3600000);

   (* change history
   hm 4. aug 2006  rev 1.0
     original version

   hm 2.10.2006   rev 1.1
     changed name of input to itod

   *)
END_FUNCTION

FUNCTION "HOUR_OF_DT" : Int   // FC188, SCL
TITLE = HOUR_OF_DT
{ S7_Optimized_Access := 'FALSE' }
AUTHOR : oscat
FAMILY : TIDT
NAME : H_DT
VERSION : 1.0
// HOUR_OF_DT returns the current hour (hour of the day) of a DT variable
   VAR_INPUT
      XDT : Date_And_Time;
      _XDT AT XDT : Array[0..7] of Byte;
   END_VAR
BEGIN


   #HOUR_OF_DT := BCD16_TO_INT(#_XDT[3]); 

   (* 
       original code:
       HOUR_OF_DT := DWORD_TO_INT((DT_TO_DWORD(XDT) MOD 86400)/3600);
   *)

   (* revision history
   hm      6.9.2008    rev 1.0
       original version


   *)
END_FUNCTION

FUNCTION "HOUR_TO_TIME" : Time   // FC189, SCL
TITLE = HOUR_TO_TIME
{ S7_Optimized_Access := 'FALSE' }
AUTHOR : hugo
FAMILY : TIDT
NAME : H2TI
VERSION : 1.2
// converts an amount of hours in real to time
   VAR_INPUT
      IN : Real;
   END_VAR
BEGIN


   #HOUR_TO_TIME := T_CONV(REAL_TO_DINT(#IN * 3600000));


   (* revision history
   hm      4. aug 2006 rev 1.0
       original version

   hm  14. mar. 2008   rev 1.1
       rounded the input after the last digit

   hm  24. feb. 2009   rev 1.2
       changed input to IN
   *)
END_FUNCTION

FUNCTION "HOUR_TO_TOD" : Time_Of_Day   // FC190, SCL
TITLE = HOUR_TO_TOD
{ S7_Optimized_Access := 'FALSE' }
AUTHOR : hugo
FAMILY : TIDT
NAME : H2TOD
VERSION : 1.1
// converts an amount of hours in real to time of day
   VAR_INPUT
      input : Real;
   END_VAR
BEGIN


     #HOUR_TO_TOD := T_CONV(REAL_TO_DINT(#input * 3600000));

   (* revision history
   hm      4. aug 2006 rev 1.0
       original version

   hm      14. mar 2008    rev 1.1
       rounded the input after the last digit

   *)
END_FUNCTION

FUNCTION "JD2000" : Real   // FC191, SCL
TITLE = JD2000
{ S7_Optimized_Access := 'FALSE' }
AUTHOR : hugo
FAMILY : TIDT
NAME : JD2000
VERSION : 1.0
// JULIAN calculates the astronomic julian date.
// 
// uses: DT_DINT [FC400]
//       DT_DATE [FC6] 
//       DT_TOD [FC8]
   VAR_INPUT
      DTI : Date_And_Time;
   END_VAR
   VAR_TEMP
      tDTI : Date_And_Time;
   END_VAR
BEGIN


   #tDTI := #DTI;
   #JD2000 := DINT_TO_REAL("DT_DINT"(#tDTI) - 946728000) / 86400.0;



   (* revision histroy
   hm  15. jul. 2008   rev 1.0
       original release


   *)
END_FUNCTION

FUNCTION "LEAP_DAY" : Bool   // FC192, SCL
TITLE = LEAP_DAY
{ S7_Optimized_Access := 'FALSE' }
AUTHOR : hugo
FAMILY : TIDT
NAME : LEAPDAY
VERSION : 1.2
// leap_day is true if the tested day is a leap day (29. of february).  
//   
// uses:  DATE_DINT (FC405)
   VAR_INPUT
      IDATE : Date;
   END_VAR
BEGIN


   #LEAP_DAY := "DATE_DINT"(#IDATE) MOD 126230400 = 68169600;


   (* change history

   hm  15. jun. 2008 rev 1.0
     original version

   hm  7. oct. 2008  rev 1.1
     changed function month to month_of_date

   hm  24. jan. 2011 rev 1.2
     improved performance
   *)
END_FUNCTION

FUNCTION "LEAP_OF_DATE" : Bool   // FC193, SCL
TITLE = LEAP_OF_DATE
{ S7_Optimized_Access := 'FALSE' }
AUTHOR : hugo
FAMILY : TIDT
NAME : LEAPODAT
VERSION : 1.3
// leap_year is true if the tested year is a leap year  
// 
// uses: DATE_DINT [FC405]
   VAR_INPUT
      idate : Date;
   END_VAR
BEGIN


   #LEAP_OF_DATE := SHL(IN:=DINT_TO_DWORD((("DATE_DINT"(#idate) + 43200) / 31557600)),N:=30) = 16#80000000;


   (* change history

   2.10.2006   rev 1.1
   the function now calls leap_year to accomodate further accuracy.
   the function now works for any year from 1970 to 2100

   8. jan 2008   rev 1.2
     improved code for better performance

   28. jan. 2011 rev 1.3
     improved performance
   *)
END_FUNCTION

FUNCTION "LEAP_YEAR" : Bool   // FC194, SCL
TITLE = LEAP_YEAR
{ S7_Optimized_Access := 'FALSE' }
AUTHOR : hugo
FAMILY : TIDT
NAME : LEAPY
VERSION : 1.1
// leap_year is true if the tested year is a leap year
   VAR_INPUT
      yr : Int;
   END_VAR
BEGIN


   IF #yr MOD 400 = 0 THEN #LEAP_YEAR := TRUE;
   ELSIF #yr MOD 100 = 0 THEN #LEAP_YEAR := FALSE;
   ELSIF #yr MOD 4 =0 THEN #LEAP_YEAR := TRUE;
   ELSE #LEAP_YEAR := FALSE;
   END_IF;


   (* change history

   2.10.2006       changes to rev 1.1
   the function now works for any year from 1970 up to 2100

   *)
END_FUNCTION

FUNCTION "LTIME_TO_UTC" : Date_And_Time   // FC196, SCL
TITLE = LTIME_TO_UTC
{ S7_Optimized_Access := 'FALSE' }
AUTHOR : hugo
FAMILY : TIDT
NAME : LT2UTC
VERSION : 1.7
// LTIME_TO_UTC calculates UTC (World Time) from a local time LTIME. utc is calculated by subtracting Time_Zone_Offset from ltime and if dst it true subtracting an additional hour from ltime.
// 
// uses: DINT_DT [FC399]
//       D_TOD_DT [FC3] 
//       DT_DINT [FC400]
//       DT_DATE [FC6] 
//       DT_TOD [FC8]
   VAR_INPUT
      LTIME : Date_And_Time;
      DST : Bool;
      TIME_ZONE_OFFSET : Int;
   END_VAR
   VAR_TEMP
      tLtime : Date_And_Time;
      tLTIME_TO_UTC : Date_And_Time;
   END_VAR
BEGIN


   #tLTIME_TO_UTC := #LTIME_TO_UTC;
   #tLtime:= #LTIME;

   #tLTIME_TO_UTC := "DINT_DT"("DT_DINT"(#tLtime) - INT_TO_DINT(#TIME_ZONE_OFFSET)*60);
   IF #DST THEN #tLTIME_TO_UTC := #tLTIME_TO_UTC T_SUB T#1h; END_IF;

   #LTIME_TO_UTC := #tLTIME_TO_UTC;

   (* revision history
   hm 5.7.2007  rev 1.0  
    original version

   hm 5.11.2007  rev 1.1
    replaced literal constant with variable because of error in möller ecp4 compiler

   hm 12.nov 2007 rev 1.2
    changed Type of time_zone_offset from time to int to allow for time zones with negative offset

   hm 8. dec 2007 rev 1.3
    corrected a problem with time_zone_offset

   hm 14. oct. 2008 rev 1.4
    changed time_zone_offset from int to real to allow for half hour offset

